// TIA Portal project "ProjectTest" (V15.1)

(* hardware
DEVICE "S7-1200 station_1"  S7-1200 Station
   slot 0: "Rack_0"  S7-1200 Rack  Rack  V1.0
   slot 1: "PLC_1"  CPU 1214C DC/DC/DC  6ES7 214-1AG40-0XB0  V4.2
DEVICE "HMI_1"  KTP900 Basic PN
   slot 0: "HMI_1"  KTP900 Basic PN  6AV2 123-2JB03-0AX0  15.1.0.0
   slot 1: "HMI_RT_1"  KTP900 Basic PN  6AV2 123-2JB03-0AX0  15.1.0.0
   slot 5: "HMI_1.IE_CP_1"  PROFINET Interface  15.0.1.0
      slot 1: "PROFINET Interface_1"  PROFINET Interface
         slot 1: "Port_1"  Port
DEVICE "S71500/ET200MP station_1"  S7-1500 station
   slot 0: "Rail_0"  Rack  6ES7 590-1***0-0AA0
   slot 1: "PLC_2"  CPU 1513-1 PN  6ES7 513-1AL02-0AB0  V2.6
      slot 3: "CPU display_1"  6ES7591-1AA00-0AA0
DEVICE "HMI_2"  KTP900 Basic PN
   slot 0: "HMI_2"  KTP900 Basic PN  6AV2 123-2JB03-0AX0  15.1.0.0
   slot 1: "HMI_RT_2"  KTP900 Basic PN  6AV2 123-2JB03-0AX0  15.1.0.0
   slot 5: "HMI_2.IE_CP_1"  PROFINET Interface  15.0.1.0
      slot 1: "PROFINET Interface_1"  PROFINET Interface
         slot 1: "Port_1"  Port
*)

// ===== PLC "PLC_1"  CPU 1214C DC/DC/DC =====

VAR_GLOBAL   // PLC tag table "Default tag table"
   "System_Byte" AT %MB1 : Byte;
   "FirstScan" AT %M1.0 : Bool;
   "DiagStatusUpdate" AT %M1.1 : Bool;
   "AlwaysTRUE" AT %M1.2 : Bool;
   "AlwaysFALSE" AT %M1.3 : Bool;
   "Clock_Byte" AT %MB0 : Byte;
   "Clock_10Hz" AT %M0.0 : Bool;
   "Clock_5Hz" AT %M0.1 : Bool;
   "Clock_2.5Hz" AT %M0.2 : Bool;
   "Clock_2Hz" AT %M0.3 : Bool;
   "Clock_1.25Hz" AT %M0.4 : Bool;
   "Clock_1Hz" AT %M0.5 : Bool;
   "Clock_0.625Hz" AT %M0.6 : Bool;
   "Clock_0.5Hz" AT %M0.7 : Bool;
   "puls" AT %M2.0 : Bool;
END_VAR

VAR_GLOBAL   // PLC tag table "Tags_DI"
   "Pompa1" AT %Q0.0 : Bool;
   "Pompa2" AT %Q0.1 : Bool;
   "Vana Consum" AT %Q0.2 : Bool;
   "Buton pompa1" AT %I0.0 : Bool;
   "Buton Pompa2" AT %I0.1 : Bool;
   "Buton Vana" AT %I0.2 : Bool;
   "Resetare Contor1" AT %I0.3 : Bool;
   "Resetare Contor2" AT %I0.4 : Bool;
   "Indicatie Pompa1" AT %I0.5 : Bool;
   "Indicatie Pompa2" AT %I0.6 : Bool;
   "Indicatie mod" AT %I0.7 : Bool;
END_VAR

DATA_BLOCK "Bazin"   // DB1
{ S7_Optimized_Access := 'TRUE' }
VERSION : 0.1
   VAR
      Nivel : Real;
      "Vana golire" : Bool := false;
      "Debit golire" : Int := 10;
      Cheie : Int := 1;
      Stare_rising_edge : Bool;
   END_VAR
BEGIN
END_DATA_BLOCK

DATA_BLOCK "Pompa_1"   // DB2
{ S7_Optimized_Access := 'TRUE' }
VERSION : 0.1
   VAR
      Stare : Bool;
      Capacitate : Real := 15.0;
      "Mod" : Int;
      Contor : UInt;
      Stare_rising_edge_bazin : Bool;
      Reset : Bool;
      add_15l : Real := 15.0;
      Stare_rising_edge_pompa : Bool;
   END_VAR
BEGIN
END_DATA_BLOCK

DATA_BLOCK "Pompa_2"   // DB3
{ S7_Optimized_Access := 'TRUE' }
VERSION : 0.1
   VAR
      Stare : Bool;
      Capacitate : Real := 15.0;
      "Mod" : Int;
      Contor : UInt;
      Stare_rising_edge_bazin : Bool;
      Reset : Bool;
      add_15l : Real := 15.0;
      State_rising_edge_pompa : Bool;
   END_VAR
BEGIN
END_DATA_BLOCK

DATA_BLOCK "Adauga  15L la bazin_DB"   // DB4
{ S7_Optimized_Access := 'TRUE' }
VERSION : 0.1
// stored: InstanceOfName Adauga 15L la bazin
"Adauga  15L la bazin"
BEGIN
END_DATA_BLOCK

DATA_BLOCK "Adauga  15L la bazin_DB_1"   // DB5
{ S7_Optimized_Access := 'TRUE' }
VERSION : 0.1
// stored: InstanceOfName Adauga 15L la bazin
"Adauga  15L la bazin"
BEGIN
END_DATA_BLOCK

DATA_BLOCK "Adauga  15L la bazin_DB_2"   // DB6
{ S7_Optimized_Access := 'TRUE' }
VERSION : 0.1
// stored: InstanceOfName Adauga 15L la bazin
"Adauga  15L la bazin"
BEGIN
END_DATA_BLOCK

DATA_BLOCK "Adauga  15L la bazin_DB_3"   // DB7
{ S7_Optimized_Access := 'TRUE' }
VERSION : 0.1
// stored: InstanceOfName Adauga 15L la bazin
"Adauga  15L la bazin"
BEGIN
END_DATA_BLOCK

DATA_BLOCK "Adauga  15L la bazin_DB_4"   // DB8
{ S7_Optimized_Access := 'TRUE' }
VERSION : 0.1
// stored: InstanceOfName Adauga 15L la bazin
"Adauga  15L la bazin"
BEGIN
END_DATA_BLOCK

DATA_BLOCK "Adauga  15L la bazin_DB_5"   // DB9
{ S7_Optimized_Access := 'TRUE' }
VERSION : 0.1
// stored: InstanceOfName Adauga 15L la bazin
"Adauga  15L la bazin"
BEGIN
END_DATA_BLOCK

DATA_BLOCK "pompa convertizor_DB"   // DB10
{ S7_Optimized_Access := 'TRUE' }
VERSION : 0.1
// stored: InstanceOfName pompa convertizor
"pompa convertizor"
BEGIN
END_DATA_BLOCK

DATA_BLOCK "pompaconvertizor variabile"   // DB11
{ S7_Optimized_Access := 'TRUE' }
VERSION : 0.1
   VAR
      "int pid" : Real;
      disponibil : Bool;
      "mod fct" : Bool;
      fault : Bool;
      ESD : Bool;
      b_start : Bool;
      B_stop : Bool;
      "viteza impusa" : Real;
      start_auto : Bool;
      "out debit" : Real;
      "cmd pmp" : Bool;
      puls_pmp_conv : Bool;
   END_VAR
BEGIN
END_DATA_BLOCK

DATA_BLOCK "pid db"   // DB13
{ S7_Optimized_Access := 'TRUE' }
VERSION : 0.1
   VAR
      setpoint : Real;
      input : Real;
      output : Real;
   END_VAR
BEGIN
END_DATA_BLOCK

FUNCTION_BLOCK "Adauga  15L la bazin"   // FB1, LAD
{ S7_Optimized_Access := 'TRUE' }
VERSION : 0.1
   VAR_INPUT
      Input_2 : Bool;
   END_VAR
   VAR_TEMP
      clock_rising_edge : Bool;
   END_VAR
   VAR_TEMP   // added for the SCL form of the ladder/FBD networks
      _w1 : Bool;
      _w2 : Bool;
   END_VAR
BEGIN

REGION Network 1
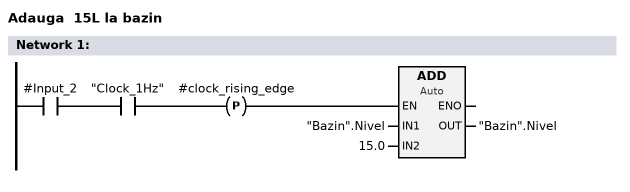
   RUNG wire#powerrail
      Contact( #Input_2 )
      Contact( "Clock_1Hz" )
      P_Trig( #clock_rising_edge )
      Add(in1 := "Bazin".Nivel, in2 := 15.0, out => "Bazin".Nivel)
   END_RUNG
   // the same network as SCL:
   #_w1 := #Input_2 AND "Clock_1Hz";
   #_w2 := #_w1 AND NOT #clock_rising_edge;   // rising edge
   #clock_rising_edge := #_w1;
   IF #_w2 THEN "Bazin".Nivel := "Bazin".Nivel + 15.0; END_IF;
END_REGION
END_FUNCTION_BLOCK

FUNCTION_BLOCK "pompa convertizor"   // FB2, LAD
{ S7_Optimized_Access := 'TRUE' }
VERSION : 0.1
   VAR_INPUT
      int_pid : Real;
      disponibil : Bool;
      mad_fct : Bool;
      fault : Bool;
      ESD : Bool;
      B_start_manual : Bool;
      B_stop_manual : Bool;
      viteza_impusa_manual : Real;
      start_auto : Bool;
   END_VAR
   VAR_OUTPUT
      out_debit : Real;
      cmd_pompa : Bool;
   END_VAR
   VAR
      reg_auto : Bool;
      reg_man : Bool;
   END_VAR
BEGIN

REGION Network 1: selctare regim auto
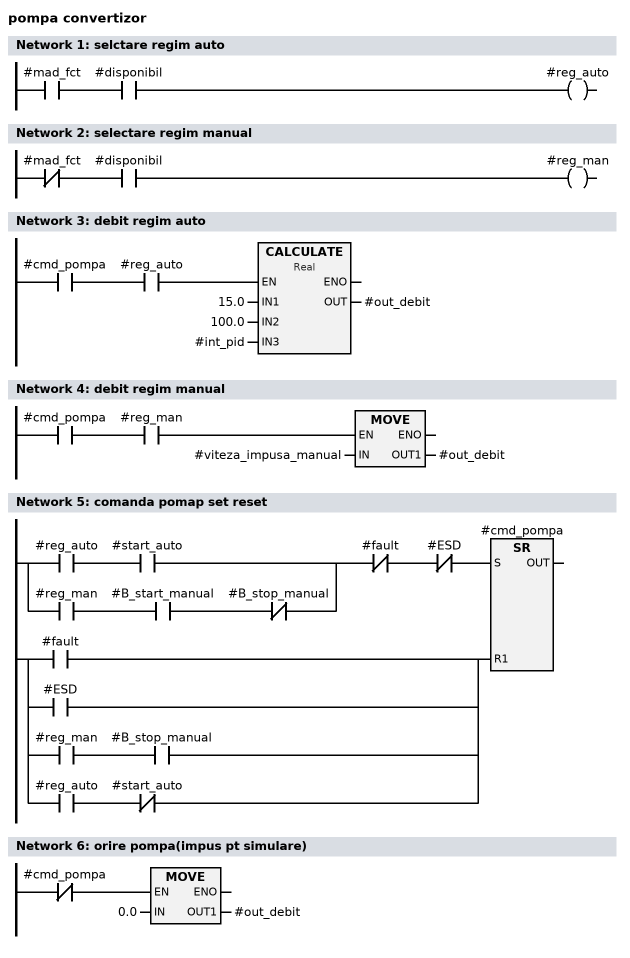
   RUNG wire#powerrail
      Contact( #mad_fct )
      Contact( #disponibil )
      Coil( #reg_auto )
   END_RUNG
   // the same network as SCL:
   #reg_auto := #mad_fct AND #disponibil;
END_REGION

REGION Network 2: selectare regim manual
   RUNG wire#powerrail
      I_Contact( #mad_fct )
      Contact( #disponibil )
      Coil( #reg_man )
   END_RUNG
   // the same network as SCL:
   #reg_man := NOT #mad_fct AND #disponibil;
END_REGION

REGION Network 3: debit regim auto
   RUNG wire#powerrail
      Contact( #cmd_pompa )
      Contact( #reg_auto )
      { S7_Templates := "SrcType := Real"; S7_Expression := "IN1 * IN3 / IN2" } Calculate(in1 := 15.0, in2 := 100.0, in3 := #int_pid, out => #out_debit)
   END_RUNG
   // the same network as SCL:
   IF #cmd_pompa AND #reg_auto THEN #out_debit := 15.0 * #int_pid / 100.0; END_IF;
END_REGION

REGION Network 4: debit regim manual
   RUNG wire#powerrail
      Contact( #cmd_pompa )
      Contact( #reg_man )
      Move(in := #viteza_impusa_manual, out1 => #out_debit)
   END_RUNG
   // the same network as SCL:
   IF #cmd_pompa AND #reg_man THEN #out_debit := #viteza_impusa_manual; END_IF;
END_REGION

REGION Network 5: comanda pomap set reset
   RUNG wire#powerrail
      Contact( #reg_auto )
      Contact( #start_auto )
      wire#w1
      I_Contact( #fault )
      I_Contact( #ESD )
      S_SR(operand := #cmd_pompa, r1 := wire#w2)
   END_RUNG
   RUNG wire#powerrail
      Contact( #reg_man )
      Contact( #B_start_manual )
      I_Contact( #B_stop_manual )
   END_RUNG wire#w1
   RUNG wire#powerrail
      Contact( #fault )
   END_RUNG wire#w2
   RUNG wire#powerrail
      Contact( #ESD )
   END_RUNG wire#w2
   RUNG wire#powerrail
      Contact( #reg_man )
      Contact( #B_stop_manual )
   END_RUNG wire#w2
   RUNG wire#powerrail
      Contact( #reg_auto )
      I_Contact( #start_auto )
   END_RUNG wire#w2
   // the same network as SCL:
   IF ((#reg_auto AND #start_auto) OR (#reg_man AND #B_start_manual AND NOT #B_stop_manual)) AND NOT #fault AND NOT #ESD THEN
       #cmd_pompa := TRUE;   // SR flip-flop
   END_IF;
   IF #fault OR #ESD OR (#reg_man AND #B_stop_manual) OR (#reg_auto AND NOT #start_auto) THEN
       #cmd_pompa := FALSE;
   END_IF;
END_REGION

REGION Network 6: orire pompa(impus pt simulare)
   RUNG wire#powerrail
      I_Contact( #cmd_pompa )
      Move(in := 0.0, out1 => #out_debit)
   END_RUNG
   // the same network as SCL:
   IF NOT #cmd_pompa THEN #out_debit := 0.0; END_IF;
END_REGION
END_FUNCTION_BLOCK

FUNCTION "Block_1" : Void   // FC1, LAD
{ S7_Optimized_Access := 'TRUE' }
VERSION : 0.1
   VAR_INPUT
      input1 : Bool;
   END_VAR
   VAR_TEMP
      clock_rising_edge : Bool;
   END_VAR
   VAR_TEMP   // added for the SCL form of the ladder/FBD networks
      _w1 : Bool;
      _w2 : Bool;
   END_VAR
BEGIN

REGION Network 1
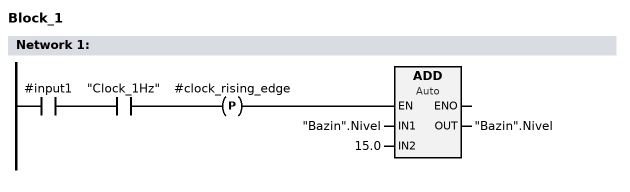
   RUNG wire#powerrail
      Contact( #input1 )
      Contact( "Clock_1Hz" )
      P_Trig( #clock_rising_edge )
      Add(in1 := "Bazin".Nivel, in2 := 15.0, out => "Bazin".Nivel)
   END_RUNG
   // the same network as SCL:
   #_w1 := #input1 AND "Clock_1Hz";
   #_w2 := #_w1 AND NOT #clock_rising_edge;   // rising edge
   #clock_rising_edge := #_w1;
   IF #_w2 THEN "Bazin".Nivel := "Bazin".Nivel + 15.0; END_IF;
END_REGION
END_FUNCTION

ORGANIZATION_BLOCK "Main"   // OB1, LAD, ProgramCycle
TITLE = "Main Program Sweep (Cycle)"
{ S7_Optimized_Access := 'TRUE' }
VERSION : 0.1
   VAR_INPUT
      Initial_Call : Bool;   // Initial call of this OB
      Remanence : Bool;   // =True, if remanent data are available
   END_VAR
   VAR_TEMP   // added for the SCL form of the ladder/FBD networks
      _w1 : Bool;
      _w2 : Bool;
      _w3 : Bool;
      _w4 : Bool;
   END_VAR
BEGIN

REGION Network 1: moduri de functionare
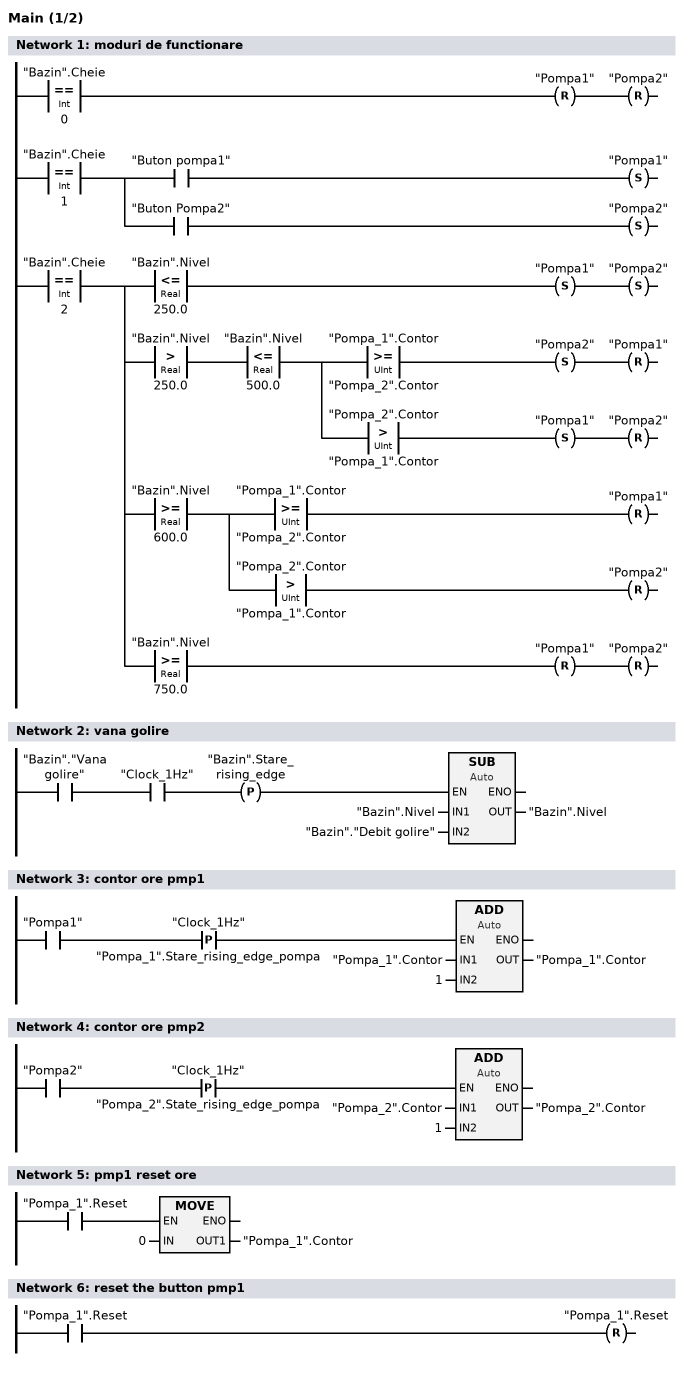
   RUNG wire#powerrail
      { S7_Templates := "SrcType := Int" } EQ_Contact(in1 := "Bazin".Cheie, in2 := 0)
      R_Coil( "Pompa1" )
      R_Coil( "Pompa2" )
   END_RUNG
   RUNG wire#powerrail
      { S7_Templates := "SrcType := Int" } EQ_Contact(in1 := "Bazin".Cheie, in2 := 1)
      wire#w1
      Contact( "Buton pompa1" )
      S_Coil( "Pompa1" )
   END_RUNG
   RUNG wire#w1
      Contact( "Buton Pompa2" )
      S_Coil( "Pompa2" )
   END_RUNG
   RUNG wire#powerrail
      { S7_Templates := "SrcType := Int" } EQ_Contact(in1 := "Bazin".Cheie, in2 := 2)
      wire#w2
      { S7_Templates := "SrcType := Real" } LE_Contact(in1 := "Bazin".Nivel, in2 := 250.0)
      S_Coil( "Pompa1" )
      S_Coil( "Pompa2" )
   END_RUNG
   RUNG wire#w2
      { S7_Templates := "SrcType := Real" } GT_Contact(in1 := "Bazin".Nivel, in2 := 250.0)
      { S7_Templates := "SrcType := Real" } LE_Contact(in1 := "Bazin".Nivel, in2 := 500.0)
      wire#w3
      { S7_Templates := "SrcType := UInt" } GE_Contact(in1 := "Pompa_1".Contor, in2 := "Pompa_2".Contor)
      S_Coil( "Pompa2" )
      R_Coil( "Pompa1" )
   END_RUNG
   RUNG wire#w3
      { S7_Templates := "SrcType := UInt" } GT_Contact(in1 := "Pompa_2".Contor, in2 := "Pompa_1".Contor)
      S_Coil( "Pompa1" )
      R_Coil( "Pompa2" )
   END_RUNG
   RUNG wire#w2
      { S7_Templates := "SrcType := Real" } GE_Contact(in1 := "Bazin".Nivel, in2 := 600.0)
      wire#w4
      { S7_Templates := "SrcType := UInt" } GE_Contact(in1 := "Pompa_1".Contor, in2 := "Pompa_2".Contor)
      R_Coil( "Pompa1" )
   END_RUNG
   RUNG wire#w4
      { S7_Templates := "SrcType := UInt" } GT_Contact(in1 := "Pompa_2".Contor, in2 := "Pompa_1".Contor)
      R_Coil( "Pompa2" )
   END_RUNG
   RUNG wire#w2
      { S7_Templates := "SrcType := Real" } GE_Contact(in1 := "Bazin".Nivel, in2 := 750.0)
      R_Coil( "Pompa1" )
      R_Coil( "Pompa2" )
   END_RUNG
   // the same network as SCL:
   IF "Bazin".Cheie = 0 THEN
       "Pompa1" := FALSE;
       "Pompa2" := FALSE;
   END_IF;
   #_w1 := "Bazin".Cheie = 1;
   IF #_w1 AND "Buton pompa1" THEN "Pompa1" := TRUE; END_IF;
   IF #_w1 AND "Buton Pompa2" THEN "Pompa2" := TRUE; END_IF;
   #_w2 := "Bazin".Cheie = 2;
   IF #_w2 AND ("Bazin".Nivel <= 250.0) THEN
       "Pompa1" := TRUE;
       "Pompa2" := TRUE;
   END_IF;
   #_w3 := #_w2 AND ("Bazin".Nivel > 250.0) AND ("Bazin".Nivel <= 500.0);
   IF #_w3 AND ("Pompa_1".Contor >= "Pompa_2".Contor) THEN
       "Pompa2" := TRUE;
       "Pompa1" := FALSE;
   END_IF;
   IF #_w3 AND ("Pompa_2".Contor > "Pompa_1".Contor) THEN
       "Pompa1" := TRUE;
       "Pompa2" := FALSE;
   END_IF;
   #_w4 := #_w2 AND ("Bazin".Nivel >= 600.0);
   IF #_w4 AND ("Pompa_1".Contor >= "Pompa_2".Contor) THEN "Pompa1" := FALSE; END_IF;
   IF #_w4 AND ("Pompa_2".Contor > "Pompa_1".Contor) THEN "Pompa2" := FALSE; END_IF;
   IF #_w2 AND ("Bazin".Nivel >= 750.0) THEN
       "Pompa1" := FALSE;
       "Pompa2" := FALSE;
   END_IF;
END_REGION

REGION Network 2: vana golire
   RUNG wire#powerrail
      Contact( "Bazin"."Vana golire" )
      Contact( "Clock_1Hz" )
      P_Trig( "Bazin".Stare_rising_edge )
      Sub(in1 := "Bazin".Nivel, in2 := "Bazin"."Debit golire", out => "Bazin".Nivel)
   END_RUNG
   // the same network as SCL:
   #_w1 := "Bazin"."Vana golire" AND "Clock_1Hz";
   #_w2 := #_w1 AND NOT "Bazin".Stare_rising_edge;   // rising edge
   "Bazin".Stare_rising_edge := #_w1;
   IF #_w2 THEN "Bazin".Nivel := "Bazin".Nivel - "Bazin"."Debit golire"; END_IF;
END_REGION

REGION Network 3: contor ore pmp1
   RUNG wire#powerrail
      Contact( "Pompa1" )
      P_Contact(operand := "Clock_1Hz", bit := "Pompa_1".Stare_rising_edge_pompa)
      Add(in1 := "Pompa_1".Contor, in2 := 1, out => "Pompa_1".Contor)
   END_RUNG
   // the same network as SCL:
   #_w1 := "Pompa1" AND "Clock_1Hz" AND NOT "Pompa_1".Stare_rising_edge_pompa;   // rising edge of "Clock_1Hz"
   "Pompa_1".Stare_rising_edge_pompa := "Clock_1Hz";
   IF #_w1 THEN "Pompa_1".Contor := "Pompa_1".Contor + 1; END_IF;
END_REGION

REGION Network 4: contor ore pmp2
   RUNG wire#powerrail
      Contact( "Pompa2" )
      P_Contact(operand := "Clock_1Hz", bit := "Pompa_2".State_rising_edge_pompa)
      Add(in1 := "Pompa_2".Contor, in2 := 1, out => "Pompa_2".Contor)
   END_RUNG
   // the same network as SCL:
   #_w1 := "Pompa2" AND "Clock_1Hz" AND NOT "Pompa_2".State_rising_edge_pompa;   // rising edge of "Clock_1Hz"
   "Pompa_2".State_rising_edge_pompa := "Clock_1Hz";
   IF #_w1 THEN "Pompa_2".Contor := "Pompa_2".Contor + 1; END_IF;
END_REGION

REGION Network 5: pmp1 reset ore
   RUNG wire#powerrail
      Contact( "Pompa_1".Reset )
      Move(in := 0, out1 => "Pompa_1".Contor)
   END_RUNG
   // the same network as SCL:
   IF "Pompa_1".Reset THEN "Pompa_1".Contor := 0; END_IF;
END_REGION

REGION Network 6: reset the button pmp1
   RUNG wire#powerrail
      Contact( "Pompa_1".Reset )
      R_Coil( "Pompa_1".Reset )
   END_RUNG
   // the same network as SCL:
   IF "Pompa_1".Reset THEN "Pompa_1".Reset := FALSE; END_IF;
END_REGION

REGION Network 7: pmp 2 reset ore
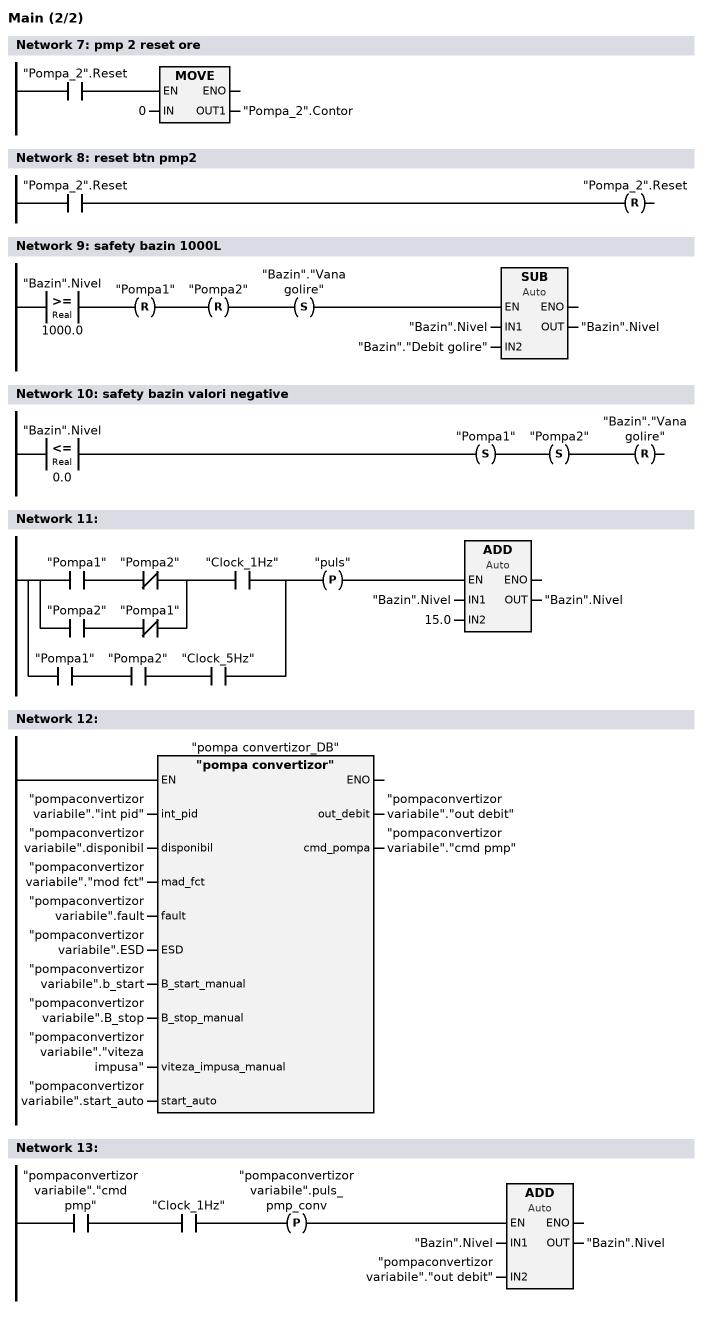
   RUNG wire#powerrail
      Contact( "Pompa_2".Reset )
      Move(in := 0, out1 => "Pompa_2".Contor)
   END_RUNG
   // the same network as SCL:
   IF "Pompa_2".Reset THEN "Pompa_2".Contor := 0; END_IF;
END_REGION

REGION Network 8: reset btn pmp2
   RUNG wire#powerrail
      Contact( "Pompa_2".Reset )
      R_Coil( "Pompa_2".Reset )
   END_RUNG
   // the same network as SCL:
   IF "Pompa_2".Reset THEN "Pompa_2".Reset := FALSE; END_IF;
END_REGION

REGION Network 9: safety bazin 1000L
   RUNG wire#powerrail
      { S7_Templates := "SrcType := Real" } GE_Contact(in1 := "Bazin".Nivel, in2 := 1000.0)
      R_Coil( "Pompa1" )
      R_Coil( "Pompa2" )
      S_Coil( "Bazin"."Vana golire" )
      Sub(in1 := "Bazin".Nivel, in2 := "Bazin"."Debit golire", out => "Bazin".Nivel)
   END_RUNG
   // the same network as SCL:
   IF "Bazin".Nivel >= 1000.0 THEN
       "Pompa1" := FALSE;
       "Pompa2" := FALSE;
       "Bazin"."Vana golire" := TRUE;
       "Bazin".Nivel := "Bazin".Nivel - "Bazin"."Debit golire";
   END_IF;
END_REGION

REGION Network 10: safety bazin valori negative
   RUNG wire#powerrail
      { S7_Templates := "SrcType := Real" } LE_Contact(in1 := "Bazin".Nivel, in2 := 0.0)
      S_Coil( "Pompa1" )
      S_Coil( "Pompa2" )
      R_Coil( "Bazin"."Vana golire" )
   END_RUNG
   // the same network as SCL:
   IF "Bazin".Nivel <= 0.0 THEN
       "Pompa1" := TRUE;
       "Pompa2" := TRUE;
       "Bazin"."Vana golire" := FALSE;
   END_IF;
END_REGION

REGION Network 11
   RUNG wire#powerrail
      Contact( "Pompa1" )
      I_Contact( "Pompa2" )
      wire#w1
      Contact( "Clock_1Hz" )
      wire#w2
      P_Trig( "puls" )
      Add(in1 := "Bazin".Nivel, in2 := 15.0, out => "Bazin".Nivel)
   END_RUNG
   RUNG wire#powerrail
      Contact( "Pompa2" )
      I_Contact( "Pompa1" )
   END_RUNG wire#w1
   RUNG wire#powerrail
      Contact( "Pompa1" )
      Contact( "Pompa2" )
      Contact( "Clock_5Hz" )
   END_RUNG wire#w2
   // the same network as SCL:
   #_w1 := ((("Pompa1" AND NOT "Pompa2") OR ("Pompa2" AND NOT "Pompa1")) AND "Clock_1Hz") OR ("Pompa1" AND "Pompa2" AND "Clock_5Hz");
   #_w2 := #_w1 AND NOT "puls";   // rising edge
   "puls" := #_w1;
   IF #_w2 THEN "Bazin".Nivel := "Bazin".Nivel + 15.0; END_IF;
END_REGION

REGION Network 12
   RUNG wire#powerrail
      "pompa convertizor_DB"(int_pid := "pompaconvertizor variabile"."int pid", disponibil := "pompaconvertizor variabile".disponibil, mad_fct := "pompaconvertizor variabile"."mod fct", fault := "pompaconvertizor variabile".fault, ESD := "pompaconvertizor variabile".ESD, B_start_manual := "pompaconvertizor variabile".b_start, B_stop_manual := "pompaconvertizor variabile".B_stop, viteza_impusa_manual := "pompaconvertizor variabile"."viteza impusa", start_auto := "pompaconvertizor variabile".start_auto, out_debit => "pompaconvertizor variabile"."out debit", cmd_pompa => "pompaconvertizor variabile"."cmd pmp")
   END_RUNG
   // the same network as SCL:
   "pompa convertizor_DB"(int_pid := "pompaconvertizor variabile"."int pid",   // "pompa convertizor"
                          disponibil := "pompaconvertizor variabile".disponibil,
                          mad_fct := "pompaconvertizor variabile"."mod fct",
                          fault := "pompaconvertizor variabile".fault,
                          ESD := "pompaconvertizor variabile".ESD,
                          B_start_manual := "pompaconvertizor variabile".b_start,
                          B_stop_manual := "pompaconvertizor variabile".B_stop,
                          viteza_impusa_manual := "pompaconvertizor variabile"."viteza impusa",
                          start_auto := "pompaconvertizor variabile".start_auto,
                          out_debit => "pompaconvertizor variabile"."out debit",
                          cmd_pompa => "pompaconvertizor variabile"."cmd pmp");
END_REGION

REGION Network 13
   RUNG wire#powerrail
      Contact( "pompaconvertizor variabile"."cmd pmp" )
      Contact( "Clock_1Hz" )
      P_Trig( "pompaconvertizor variabile".puls_pmp_conv )
      Add(in1 := "Bazin".Nivel, in2 := "pompaconvertizor variabile"."out debit", out => "Bazin".Nivel)
   END_RUNG
   // the same network as SCL:
   #_w1 := "pompaconvertizor variabile"."cmd pmp" AND "Clock_1Hz";
   #_w2 := #_w1 AND NOT "pompaconvertizor variabile".puls_pmp_conv;   // rising edge
   "pompaconvertizor variabile".puls_pmp_conv := #_w1;
   IF #_w2 THEN "Bazin".Nivel := "Bazin".Nivel + "pompaconvertizor variabile"."out debit"; END_IF;
END_REGION
END_ORGANIZATION_BLOCK

ORGANIZATION_BLOCK "pid block"   // OB30, LAD, CyclicInterrupt
{ S7_Optimized_Access := 'TRUE' }
VERSION : 0.1
   VAR_INPUT
      Initial_Call : Bool;   // Initial call of this OB
      Event_Count : Int;   // Events discarded
   END_VAR
BEGIN

REGION Network 1
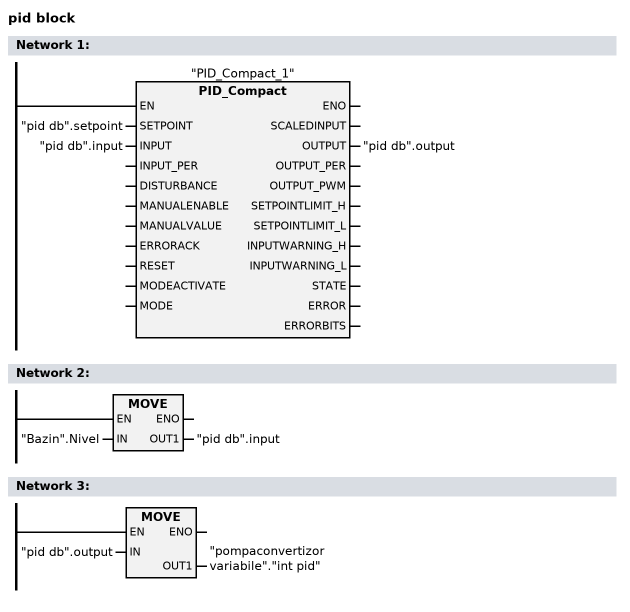
   "PID_Compact_1"(Setpoint := "pid db".setpoint, Input := "pid db".input, Output => "pid db".output);   // PID_Compact
END_REGION

REGION Network 2
   RUNG wire#powerrail
      Move(in := "Bazin".Nivel, out1 => "pid db".input)
   END_RUNG
   // the same network as SCL:
   "pid db".input := "Bazin".Nivel;
END_REGION

REGION Network 3
   RUNG wire#powerrail
      Move(in := "pid db".output, out1 => "pompaconvertizor variabile"."int pid")
   END_RUNG
   // the same network as SCL:
   "pompaconvertizor variabile"."int pid" := "pid db".output;
END_REGION
END_ORGANIZATION_BLOCK

// ===== PLC "PLC_2"  CPU 1513-1 PN =====

VAR_GLOBAL   // PLC tag table "Default tag table"
   "Clock_Byte" AT %MB0 : Byte;
   "Clock_10Hz" AT %M0.0 : Bool;
   "Clock_5Hz" AT %M0.1 : Bool;
   "Clock_2.5Hz" AT %M0.2 : Bool;
   "Clock_2Hz" AT %M0.3 : Bool;
   "Clock_1.25Hz" AT %M0.4 : Bool;
   "Clock_1Hz" AT %M0.5 : Bool;
   "Clock_0.625Hz" AT %M0.6 : Bool;
   "Clock_0.5Hz" AT %M0.7 : Bool;
END_VAR

DATA_BLOCK "@pompa convertizor_DB"   // DB1
{ S7_Optimized_Access := 'TRUE' }
VERSION : 0.1
// stored: InstanceOfName pompa convertizor
"pompa convertizor"
BEGIN
END_DATA_BLOCK

DATA_BLOCK "DB_main"   // DB2
{ S7_Optimized_Access := 'TRUE' }
VERSION : 0.1
   VAR
      nivel : Real;
      vana : Bool;
      "puls vana" : Bool;
      "debit vana" : Real;
      pmp1_puls : Bool;
      pmp2_puls : Bool;
      pmp1_contor : Int;
      pmp2_contor : Int;
      pmp1_reset : Bool;
      pmp2_reset : Bool;
      selector_fct : Int := 0;
   END_VAR
BEGIN
END_DATA_BLOCK

DATA_BLOCK "db pid"   // DB4
{ S7_Optimized_Access := 'TRUE' }
VERSION : 0.1
   VAR
      setpoint : Real;
   END_VAR
BEGIN
END_DATA_BLOCK

DATA_BLOCK "db main pmp 2"   // DB5
{ S7_Optimized_Access := 'TRUE' }
VERSION : 0.1
   VAR
      "int pid" : Real;
      disponibil : Bool;
      "mod  fct" : Bool;
      fault : Bool;
      ESD : Bool;
      b_start : Bool;
      b_stop : Bool;
      "viteza impusa" : Real;
      start_auto : Bool;
      "out debit" : Real;
      "cmd pmp 2" : Bool;
      "puls pmp conv2" : Bool;
   END_VAR
BEGIN
END_DATA_BLOCK

DATA_BLOCK "pompa convertizor_DB"   // DB6
{ S7_Optimized_Access := 'TRUE' }
VERSION : 0.1
// stored: InstanceOfName pompa convertizor
"pompa convertizor"
BEGIN
END_DATA_BLOCK

DATA_BLOCK "block fct selectare_DB"   // DB7
{ S7_Optimized_Access := 'TRUE' }
VERSION : 0.1
// stored: InstanceOfName block fct selectare
"block fct selectare"
BEGIN
END_DATA_BLOCK

DATA_BLOCK "pompaconvertizor variabile"   // DB11
{ S7_Optimized_Access := 'TRUE' }
VERSION : 0.1
   VAR
      "int pid" : Real;
      disponibil : Bool;
      "mod fct" : Bool;
      fault : Bool;
      ESD : Bool;
      b_start : Bool;
      B_stop : Bool;
      "viteza impusa" : Real;
      start_auto : Bool;
      "out debit" : Real;
      "cmd pmp" : Bool;
      puls_pmp_conv : Bool;
   END_VAR
BEGIN
END_DATA_BLOCK

FUNCTION_BLOCK "block fct selectare"   // FB1, LAD
{ S7_Optimized_Access := 'TRUE' }
VERSION : 0.1
   VAR_INPUT
      "ore fct pmp1" : Real;
      "ore fct pmp 2" : Real;
      "disp 1" : Bool;
      "disp 2" : Bool;
   END_VAR
   VAR_OUTPUT
      selector_pornire : Int;
   END_VAR
BEGIN

REGION Network 1: mod 0, nu porni nicio pompa(just do nothing ig)